               (*
               FOR #Temp_Index_i := #ServerVersion_StartNum TO #MessageLen - 1 DO   //去掉前面的8个数据，同时从0开始，所以-9
                   #SaltString[#Temp_Index_i - #ServerVersion_StartNum + 2] := #REV_Buffer[#ServerVersion_StartNum];//挑战字符串的后面N个Byte
                   #ServerVersion_StartNum := #ServerVersion_StartNum + 1;
               END_FOR;*)
           END_REGION

           REGION Client_Auth_Packet
               #Temp_NowNum := 0;
               #Client_MaxLen := DINT_TO_DWORD(#MessageMaxLen);
               // Length                            3     Byte   最后处理
               #Temp_NowNum := #Temp_NowNum +3;
               // Sequence                      1     Byte
               #SND_Buffer[#Temp_NowNum] :=SINT_TO_BYTE( DINT_TO_SINT(#CDD.Connect_Sequence + 1));
               #Temp_NowNum := #Temp_NowNum + 1;
               // CapabilityFlag               4     Byte
               #SND_Buffer[#Temp_NowNum] := #Client_CapabilityFlag.%B0;
               #Temp_NowNum := #Temp_NowNum + 1;
               #SND_Buffer[#Temp_NowNum] := #Client_CapabilityFlag.%B1;
               #Temp_NowNum := #Temp_NowNum + 1;
               #SND_Buffer[#Temp_NowNum] := #Client_CapabilityFlag.%B2;
               #Temp_NowNum := #Temp_NowNum + 1;
               #SND_Buffer[#Temp_NowNum] := #Client_CapabilityFlag.%B3;
               #Temp_NowNum := #Temp_NowNum + 1;
               // Max_Length                   4     Byte
               #SND_Buffer[#Temp_NowNum] := #Client_MaxLen.%B0;
               #Temp_NowNum := #Temp_NowNum + 1;
               #SND_Buffer[#Temp_NowNum] := #Client_MaxLen.%B1;
               #Temp_NowNum := #Temp_NowNum + 1;
               #SND_Buffer[#Temp_NowNum] := #Client_MaxLen.%B2;
               #Temp_NowNum := #Temp_NowNum + 1;
               #SND_Buffer[#Temp_NowNum] := #Client_MaxLen.%B3;
               #Temp_NowNum := #Temp_NowNum + 1;
               // CharacterSet                 1     Byte
               #SND_Buffer[#Temp_NowNum] := #CDD.Server_Character_Set;
               #Temp_NowNum := #Temp_NowNum + 1;
               // Fill Data  (16#00)          23  Byte
               FOR #Temp_Index_i := 0 TO 22 DO
                   #SND_Buffer[#Temp_NowNum + #Temp_Index_i] := b#16#00;
               END_FOR;
               #Temp_NowNum := #Temp_NowNum + 23;
               // User Name                    N    Byte    Last Character    16#00
               #Temp_StrLen := LEN(#UserName);
               FOR #Temp_Index_i := 0 TO #Temp_StrLen - 1 DO
                   #SND_Buffer[#Temp_NowNum + #Temp_Index_i] := #UserName[#Temp_Index_i + 1];
               END_FOR;
               #Temp_NowNum := #Temp_NowNum + #Temp_StrLen;
               #SND_Buffer[#Temp_NowNum] := b#16#00;
               #Temp_NowNum := #Temp_NowNum + 1;
               #SND_Buffer[#Temp_NowNum] := b#16#14;
               #Temp_NowNum := #Temp_NowNum + 1;
               // Token                              N    Byte    Last Character    16#00
               #Calc_Encryption_SHA1(IN_Str := #PassWord,
                                     TempOutStr => #Temp_SHA1);
               #Calc_Encryption_SHA1(IN_Str := #Temp_SHA1,
                                     Len:=20,
                                     TempOutStr => #Temp_SHA1_2);
               // Strg_TO_Chars(Strg := #PassWord,
               //               pChars := 0,
               //               Cnt => #Temp_SHA_Arry_Num,
               //               Chars := #Temp_SHA_Arry);
               // #Temp_SHA_Arry_Num_Int := UINT_TO_INT(#Temp_SHA_Arry_Num);

               FOR #Temp_Index_i := 0 TO 19 DO
                   #Temp_SHA_Arry[#Temp_Index_i] := #SaltString[#Temp_Index_i];
               END_FOR;
               FOR #Temp_Index_i := 20 TO 39 DO
                   #Temp_SHA_Arry[#Temp_Index_i] := #Temp_SHA1_2[#Temp_Index_i - 20];
               END_FOR;

               #Calc_Encryption_SHA1(IN_Str := #Temp_SHA_Arry,
                                     Len := 40,
                                     TempOutStr => #Temp_SHA1_3);

               FOR #Temp_Index_i := 0 TO 19 DO
                   #Token[#Temp_Index_i] := #Temp_SHA1[#Temp_Index_i] XOR #Temp_SHA1_3[#Temp_Index_i];
                   #SND_Buffer[#Temp_NowNum + #Temp_Index_i] := #Token[#Temp_Index_i];
               END_FOR;
               #Temp_NowNum := #Temp_NowNum + 20;
               #SND_Buffer[#Temp_NowNum] := b#16#00;
               #Temp_NowNum := #Temp_NowNum + 1;

               // DataBase Name           N    Byte    Last Character    16#00
               #Temp_StrLen := LEN(#DB_Name);
               FOR #Temp_Index_i := 0 TO #Temp_StrLen - 1 DO
                   #SND_Buffer[#Temp_NowNum + #Temp_Index_i] := #DB_Name[#Temp_Index_i + 1];
               END_FOR;
               #Temp_NowNum := #Temp_NowNum + #Temp_StrLen;
               #SND_Buffer[#Temp_NowNum] := b#16#00;
               #Temp_NowNum := #Temp_NowNum + 1;
               //CLIENT_PLUGIN_AUTH
               #Temp_StrLen := LEN(#CDD.CLIENT_PLUGIN_AUTH);
               FOR #Temp_Index_i := 0 TO #Temp_StrLen - 1 DO
                   #SND_Buffer[#Temp_NowNum + #Temp_Index_i] := #CDD.CLIENT_PLUGIN_AUTH[#Temp_Index_i + 1];
               END_FOR;
               #Temp_NowNum := #Temp_NowNum + #Temp_StrLen;
               #SND_Buffer[#Temp_NowNum] := b#16#00;
               #Temp_NowNum := #Temp_NowNum + 1;

               //数据长度写入前三个byte
               #Temp_Dword := DINT_TO_DWORD(INT_TO_DINT(#Temp_NowNum - 4));
               #SND_Buffer[0] := #Temp_Dword.%B0;
               #SND_Buffer[1] := #Temp_Dword.%B1;
               #SND_Buffer[2] := #Temp_Dword.%B2;
               #Step := 3;
               #NetSendLen := #Temp_NowNum;
           END_REGION

           ;

       3:  // 等待发送完成
           #NetRcv_EN := TRUE;
           #NetSend_EN := TRUE;
           IF #NetSend_Done THEN
               #NetSend_Done := FALSE;
               #NetSend_EN := FALSE;
               #Step := 4;
           END_IF;

       4:  // 等待接收数据

           IF    #NetRcv_Done  THEN
               #NetRcv_Done := FALSE;

              // #NetRcv_Len := UDINT_TO_INT(#NetRcv.RCVD_LEN);
               #NetRcv_EN := FALSE;
               #Step := 5;
           END_IF;
       5:  // 如果在等待服务器第一次连接
           IF #REV_Buffer[5]=b#16#00 AND  #NetRcv_Len >7 THEN
               #Temp_CND := TRUE;
               #NetRcv_EN := TRUE;
           END_IF;


       6:  // 申请服务器断开连接
            #SND_Buffer[0] := b#16#01;
            #SND_Buffer[1] := b#16#00;
            #SND_Buffer[2] := b#16#00;
            #SND_Buffer[3] := b#16#00;
            #SND_Buffer[4] := b#16#01;
            #NetSendEnd_EN := TRUE;
            IF #NetSendEnd_Done THEN
                #Step := 7;
            END_IF;

        7:  // 申请服务器断开连接

            #NetDiscon_EN := TRUE;
        8:
            ;
       ELSE  // Statement section ELSE
           ;
   END_CASE;


   (***********************************************************发送数据******************************************************************)
       #NetSend(REQ := #NetSend_EN,
                ID := #Net_ID,
                // DONE=>#NetSend_Done,
                LEN := INT_TO_UDINT(#NetSendLen),// INT_TO_UINT(#Temp_NowNum),
                DATA := #SND_Buffer);
       IF #NetSend.DONE THEN
           #NetSend_Done := TRUE;
       END_IF;

       #NetSendEnd(REQ := #NetSendEnd_EN,
                   ID := #Net_ID,
                   LEN := 5,
                   DONE => #NetSendEnd_Done,
                   DATA := #SND_Buffer);





   (***********************************************************断开连接******************************************************************)

   #NetDISCON(REQ:=#NetDiscon_EN AND #Timer_ON.Q ,
              ID:=#Net_ID);

   #Timer_ON(IN := NOT #Timer_OFF.Q,
             PT := t#0.5s);

   #Timer_OFF(IN := #Timer_ON.Q,
              PT := t#0.5s);




   (***********************************************************监测连接******************************************************************)
   #NetDiag(REQ := #Timer_ON.Q,
            ID := #Net_ID,
            RESULT := #TDiag_Result);
   IF  #NetDiag.ERROR THEN
       #Temp_ConnStatus := B#16#00;
   END_IF;
   IF #NetDiag.DONE THEN
       #Temp_ConnStatus := #TDiag_Result.State;
   END_IF;
   IF #Temp_ConnStatus <> B#16#04 THEN
       #Temp_CND := FALSE;
   END_IF;

   #CDD.Connect_OK := #Temp_CND;

   #Timer_Error(IN := #Connect AND NOT #Temp_CND,
                PT := t#10s);

   #Error := #Timer_Error.Q;
   #CND := #Temp_CND;
   #ConnStatus := #Temp_ConnStatus;

   (***********************************************************数据传递******************************************************************)
   #CDD.Recv_Buffer := #REV_Buffer;
   IF #NetRcv.NDR THEN
       #CDD.Recv_Done := TRUE;
       #CDD.Recv_Len := UDINT_TO_INT(#NetRcv.RCVD_LEN);
   END_IF;
END_FUNCTION_BLOCK

FUNCTION_BLOCK "uMySQL_Query"   // FB5, SCL
{ S7_Optimized_Access := 'TRUE' }
VERSION : 0.1
   VAR_INPUT
      Command : WString[2048];
      Execute : Bool;
   END_VAR
   VAR_OUTPUT
      Done : Bool;
      Busy : Bool;
      Error : Bool;
   END_VAR
   VAR_IN_OUT
      CDD : "uMySQL_CDD";
   END_VAR
   VAR
      Net_Send : TSEND;
      Net_Send_EN : Bool;
      Net_Send_Done : Bool;
      Net_Send_Len : UInt;
      Command_Len : UInt;
      Net_Recv_EN : Bool;
      Net_Recv_Done : Bool;
      Net_Recv_Len : UInt;
      Temp_Bool : Array[0..19] of Bool;
      SendBuffer : Array[0..2048] of Byte;
      RecvBuffer : Array[0..2048] of Byte;
      SendBufferWChar : Array[0..2048] of WChar;
      TRCV : TRCV;
      Function_Run : Bool;
      Timer_instance : TON_TIME;
   END_VAR
   VAR_TEMP
      Temp_Index_i : Int;
      Temp_Dword : DWord;
      Temp_word : Word;
      Temp_Num : Int;
   END_VAR
BEGIN

   IF #Execute THEN
       #Function_Run:= TRUE;
   END_IF;

   IF #Function_Run AND NOT #Temp_Bool[0] THEN
       #Temp_Bool[0] := TRUE;
       #Net_Send_EN := TRUE;
       #Command_Len := INT_TO_UINT(LEN(#Command));
       #SendBuffer[4] := B#16#03;

       Strg_TO_Chars(Strg := #Command,
                     pChars := 0,
                     Cnt => #Command_Len,
                     Chars := #SendBufferWChar);
       (*  
       FOR #Temp_Index_i := 0 TO UINT_TO_INT( #Command_Len) -1 DO
           #SendBuffer[#Temp_Index_i + 5]:=WCHAR_TO_BYTE(#SendBufferWChar[#Temp_Index_i]) ;

       END_FOR;
       #Net_Send_Len := #Command_Len + 5;
       *)
       #Net_Send_Len := 5;

       FOR #Temp_Index_i := 0 TO UINT_TO_INT(#Command_Len) - 1 DO

           #Temp_Dword := "Wchar_To_UTF8"("WChar" := #SendBufferWChar[#Temp_Index_i], Num => #Temp_Num);
           CASE #Temp_Num OF
               1:  // 如果是单字符
                   #SendBuffer[#Net_Send_Len] := #Temp_Dword.%B0;
                   #Net_Send_Len := #Net_Send_Len + 1;
               2:  // 如果是两字节
                   #SendBuffer[#Net_Send_Len] := #Temp_Dword.%B1;
                   #Net_Send_Len := #Net_Send_Len + 1;
                   #SendBuffer[#Net_Send_Len] := #Temp_Dword.%B0;
                   #Net_Send_Len := #Net_Send_Len + 1;
               ELSE  // 如果是其他情况
                   #SendBuffer[#Net_Send_Len] := #Temp_Dword.%B2;
                   #Net_Send_Len := #Net_Send_Len + 1;
                   #SendBuffer[#Net_Send_Len] := #Temp_Dword.%B1;
                   #Net_Send_Len := #Net_Send_Len + 1;
                   #SendBuffer[#Net_Send_Len] := #Temp_Dword.%B0;
                   #Net_Send_Len := #Net_Send_Len + 1;
           END_CASE;

       END_FOR;

       #Net_Send_EN := TRUE; 
                                 //数据长度写入前三个byte
                                 #Temp_Dword := DINT_TO_DWORD(INT_TO_DINT(UINT_TO_INT(#Net_Send_Len) - 4));
                                 #SendBuffer[0] := #Temp_Dword.%B0;
                                 #SendBuffer[1] := #Temp_Dword.%B1;
                                 #SendBuffer[2] := #Temp_Dword.%B2;
                             END_IF;


   IF NOT #Function_Run THEN
       #Temp_Bool[0] := FALSE;
       #Net_Recv_Len := 0;
       #Net_Recv_Done := FALSE;
       #Net_Send_EN := FALSE;
       #Net_Recv_EN := FALSE;
       #Error := FALSE;
       #Done := FALSE;
   END_IF;


   #Net_Send(REQ:=#Net_Send_EN,
             ID:=#CDD.Connect_ID,
             LEN:=#Net_Send_Len,
             DONE=>#Net_Send_Done,
             DATA:=#SendBuffer);

   IF #Net_Send.DONE OR #Net_Send.ERROR THEN
       #Net_Send_EN := FALSE;
       #Function_Run := FALSE;
       IF #Net_Send.ERROR THEN
           #Error := TRUE;
       END_IF;
   END_IF;


   IF #CDD.Recv_Done AND #Function_Run THEN
       #Temp_word.%B0 := #CDD.Recv_Buffer[0];
       #Temp_word.%B1 := #CDD.Recv_Buffer[1];
       IF #CDD.Recv_Len = (WORD_TO_INT(#Temp_word)+4) THEN

           CASE BYTE_TO_INT(#CDD.Recv_Buffer[4]) OF
               0:
                   #Done := TRUE;
               255:  // Statement section case 2 to 4
                   #Error := TRUE;
               ELSE  // Statement section ELSE
                   ;
           END_CASE; //通过返回的数据判断是否执行成功
       ELSE
           #Error := TRUE;//如果接收的数据长度和范围数据中给定的不同则认定是通信错误
       END_IF;
       #CDD.Recv_Done := FALSE;
   END_IF;


   #Timer_instance(IN:=#Function_Run AND ( NOT #Done),
                   PT:=t#1s  );
   IF #Timer_instance.Q THEN    //如果命令执行超时，也认为是故障
       #Error := TRUE;
   END_IF;

   IF #Error THEN
       #Function_Run := FALSE;
   END_IF;
   IF #Done THEN
       #Function_Run := FALSE;
   END_IF;
END_FUNCTION_BLOCK

FUNCTION_BLOCK "Calc_Encryption_SHA1"   // FB6, SCL
{ S7_Optimized_Access := 'FALSE' }
VERSION : 0.1
   VAR_INPUT
      IN_Str : Variant;
      Len : Int;
   END_VAR
   VAR_OUTPUT
      TempOutStr : Array[0..19] of Byte;
      Encrption AT TempOutStr : Array[0..4] of DWord;
   END_VAR
   VAR_TEMP
      "A" : DWord;
      "B" : DWord;
      C : DWord;
      D : DWord;
      "E" : DWord;
      Length : Int;
      Lenth_Uint : UInt;
      MessageBlock : Array[0..63] of Byte;
      MessageBlock_DWORD AT MessageBlock : Array[0..15] of DWord;
      W : Array[0..79] of DWord;
      Index_i : Int;
      temp : DWord;
      Temp_Str : String;
      Temp_Array : Array[0..446] of Byte;
   END_VAR
   VAR CONSTANT
      K0 : DWord := 16#5A827999;   // K0计算常量
      K1 : DWord := 16#6ED9EBA1;   // K1计算常量
      K2 : DWord := 16#8F1BBCDC;   // K2计算常量
      K3 : DWord := 16#CA62C1D6;   // K3计算常量
      Const_A : DWord := 16#67452301;   // 链接变量A
      Const_B : DWord := 16#EFCDAB89;   // 链接变量B
      Const_C : DWord := 16#98BADCFE;   // 链接变量C
      Const_D : DWord := 16#10325476;   // 链接变量D
      Const_E : DWord := 16#C3D2E1F0;   // 链接变量E
   END_VAR
BEGIN
   (***************************************************数据初始化******************************************************)
   #A := #Const_A;
   #B := #Const_B;
   #C := #Const_C;
   #D := #Const_D;
   #E := #Const_E;
   //#Length := LEN(#IN_Str);
   FILL_BLK(IN := B#16#00,  COUNT := 64,  OUT => #MessageBlock[0]);
   FILL_BLK(IN := DW#16#000000000,   COUNT := 80,  OUT => #W[0]);




   (*************************************************填充/准备数据****************************************************)
   IF TypeOf(#IN_Str) =String THEN
       //如果是字符串
       VariantGet(SRC:=#IN_Str,
                  DST=>#Temp_Str);
       #Length := LEN(#Temp_Str);

       Strg_TO_Chars(Strg :=#Temp_Str ,
                     pChars := 0,
                     Cnt => #Lenth_Uint,
                     Chars := #MessageBlock);   //填充客户输入字符
   ELSE
       IF IS_ARRAY(#IN_Str) THEN
          // #Length:=UDINT_TO_INT(CountOfElements(#IN_Str)) ;
           #Length := #Len;
           VariantGet(SRC:=#IN_Str,     DST=>#Temp_Array);
           MOVE_BLK(IN := #Temp_Array[0],  COUNT :=INT_TO_UINT( #Length),  OUT => #MessageBlock[0]);
       END_IF;
     ;
   END_IF;
   (*********************************************输入数据安全检测****************************************************)
   IF (#Length = 0) OR (#Length > 56) THEN
       RETURN;
   END_IF;

   #MessageBlock[#Length] := B#16#80;   //后一位填1，其他全为0
   #MessageBlock_DWORD[14] :=DW#16#00000000;          //填充数据长度高位
   #MessageBlock_DWORD[15] := DINT_TO_DWORD(#Length * 8);//填充数据长度低位
   MOVE_BLK(IN := #MessageBlock_DWORD[0],  COUNT := 16,  OUT => #W[0]);
   FOR #Index_i := 16 TO 79 DO
       #W[#Index_i] := ROL(N := 1, IN := (#W[#Index_i - 3] XOR #W[#Index_i - 8] XOR #W[#Index_i - 14] XOR #W[#Index_i - 16]));
   END_FOR;
   (*************************************************计算过程****************************************************)
   FOR #Index_i := 0 TO 19 DO
       #temp := ROL(IN := #A, N := 5) + ((#B AND #C) OR (NOT (#B) AND #D)) + #E + #W[#Index_i] + #K0;
       #E := #D;
       #D := #C;
       #C := ROL(IN := #B, N := 30);
       #B := #A;
       #A := #temp;
   END_FOR;

   FOR #Index_i := 20 TO 39 DO
       #temp := ROL(IN := #A, N := 5) + (#B XOR #C XOR #D) + #E + #W[#Index_i] + #K1;
       #E := #D;
       #D := #C;
       #C := ROL(N := 30, IN := #B);
       #B := #A;
       #A := #temp;
   END_FOR;

   FOR #Index_i := 40 TO 59 DO
       #temp := ROL(N := 5, IN := #A) + ((#B AND #C) OR (#B AND #D) OR (#C AND #D)) + #E + #W[#Index_i] + #K2;
       #E := #D;
       #D := #C;
       #C := ROL(N := 30, IN := #B);
       #B := #A;
       #A := #temp;
   END_FOR;

   FOR #Index_i := 60 TO 79 DO
       #temp := ROL(N := 5, IN := #A) + (#B XOR #C XOR #D) + #E + #W[#Index_i] + #K3;
       #E := #D;
       #D := #C;
       #C := ROL(N := 30, IN := #B);
       #B := #A;
       #A := #temp;
   END_FOR;

   #Encrption[0] := #Const_A + #A;
   #Encrption[1] := #Const_B+ #B;
   #Encrption[2] := #Const_C + #C;
   #Encrption[3] := #Const_D + #D;
   #Encrption[4] := #Const_E + #E;
END_FUNCTION_BLOCK

FUNCTION_BLOCK "uMySQL_Use"   // FB8, SCL
{ S7_Optimized_Access := 'TRUE' }
VERSION : 0.1
   VAR_INPUT
      DB_Name : WString[2048];
      Execute : Bool;
   END_VAR
   VAR_OUTPUT
      Done : Bool;
      Busy : Bool;
      Error : Bool;
   END_VAR
   VAR_IN_OUT
      CDD : "uMySQL_CDD";
   END_VAR
   VAR
      Net_Send : TSEND;
      Net_Send_EN : Bool;
      Net_Send_Done : Bool;
      Net_Send_Len : UInt;
      Command_Len : UInt;
      Net_Recv_EN : Bool;
      Net_Recv_Done : Bool;
      Net_Recv_Len : UInt;
      Temp_Bool : Array[0..19] of Bool;
      SendBuffer : Array[0..2048] of Byte;
      RecvBuffer : Array[0..2048] of Byte;
      SendBufferWChar : Array[0..2048] of WChar;
      TRCV : TRCV;
      Function_Run : Bool;
      Timer_instance : TON_TIME;
   END_VAR
   VAR_TEMP
      Temp_Index_i : Int;
      Temp_Dword : DWord;
      Temp_word : Word;
   END_VAR
BEGIN

   IF #Execute THEN
       #Function_Run:= TRUE;
   END_IF;

   IF #Function_Run AND NOT #Temp_Bool[0] THEN
       #Temp_Bool[0] := TRUE;
       #Net_Send_EN := TRUE;
       #Command_Len := INT_TO_UINT(LEN(#DB_Name));
       #SendBuffer[4] := B#16#02;

       Strg_TO_Chars(Strg := #DB_Name,
                     pChars := 0,
                     Cnt => #Command_Len,
                     Chars := #SendBufferWChar);

       FOR #Temp_Index_i := 0 TO UINT_TO_INT(#Command_Len) - 1 DO
           #SendBuffer[#Temp_Index_i + 5] := WCHAR_TO_BYTE(#SendBufferWChar[#Temp_Index_i]);
       END_FOR;
       #Net_Send_Len := #Command_Len + 5;
       #Net_Send_EN := TRUE;
       //数据长度写入前三个byte
       #Temp_Dword := DINT_TO_DWORD(INT_TO_DINT(UINT_TO_INT(#Net_Send_Len) - 4));
       #SendBuffer[0] := #Temp_Dword.%B0;
       #SendBuffer[1] := #Temp_Dword.%B1;
       #SendBuffer[2] := #Temp_Dword.%B2;
   END_IF;


   IF NOT #Function_Run THEN
       #Temp_Bool[0] := FALSE;
       #Net_Recv_Len := 0;
       #Net_Recv_Done := FALSE;
       #Net_Send_EN := FALSE;
       #Net_Recv_EN := FALSE;
       #Error := FALSE;
       #Done := FALSE;
   END_IF;


   #Net_Send(REQ:=#Net_Send_EN,
             ID:=#CDD.Connect_ID,
             LEN:=#Net_Send_Len,
             DONE=>#Net_Send_Done,
             DATA:=#SendBuffer);

   IF #Net_Send.DONE OR #Net_Send.ERROR THEN
       #Net_Send_EN := FALSE;
       #Function_Run := FALSE;
       IF #Net_Send.ERROR THEN
           #Error := TRUE;
       END_IF;
   END_IF;


   IF #CDD.Recv_Done AND #Function_Run THEN
       #Temp_word.%B0 := #CDD.Recv_Buffer[0];
       #Temp_word.%B1 := #CDD.Recv_Buffer[1];
       IF #CDD.Recv_Len = (WORD_TO_INT(#Temp_word)+4) THEN

           CASE BYTE_TO_INT(#CDD.Recv_Buffer[4]) OF
               0:
                   #Done := TRUE;
               255:  // Statement section case 2 to 4
                   #Error := TRUE;
               ELSE  // Statement section ELSE
                   ;
           END_CASE; //通过返回的数据判断是否执行成功
       ELSE
           #Error := TRUE;//如果接收的数据长度和范围数据中给定的不同则认定是通信错误
       END_IF;
       #CDD.Recv_Done := FALSE;
   END_IF;

   #Timer_instance(IN:=#Function_Run AND ( NOT #Done),
                   PT:=t#1s  );
   IF #Timer_instance.Q THEN    //如果命令执行超时，也认为是故障
       #Error := TRUE;
   END_IF;

   IF #Error THEN
       #Function_Run := FALSE;
   END_IF;
   IF #Done THEN
       #Function_Run := FALSE;
   END_IF;
END_FUNCTION_BLOCK

FUNCTION_BLOCK "uMySQL_Command"   // FB909, SCL
{ S7_Optimized_Access := 'TRUE' }
VERSION : 0.1
   VAR
      Command : WString[2048];
   END_VAR
   VAR_TEMP
      TempStr : WString;
   END_VAR
BEGIN
   "数据库字符串"."wstring" :=WSTRING#'INSERT INTO rb001011(Addr,temp_LF,temp_RF,temp_LB,temp_RB,Distance_L,Distance_R,';
   "数据库字符串"."wstring" := CONCAT(IN1 := "数据库字符串"."wstring", IN2 := WSTRING#'Motor_Current,Motor_Freq,Motor_Power,Motor_Eng,Motor_Runhours,');
   "数据库字符串"."wstring" := CONCAT(IN1 := "数据库字符串"."wstring", IN2 := WSTRING#'EN_Temp,EN_RH,temp_Ruber,');
   "数据库字符串"."wstring" := CONCAT(IN1 := "数据库字符串"."wstring", IN2 := WSTRING#'Motor_Ready,Motor_Running,Motor_Fault,');
   "数据库字符串"."wstring" := CONCAT(IN1 := "数据库字符串"."wstring", IN2 := WSTRING#'SerialNum,Operator');
   "数据库字符串"."wstring" := CONCAT(IN1 := "数据库字符串"."wstring", IN2 := WSTRING#')VALUES(');

   "数据库字符串"."wstring" := CONCAT(IN1 := "数据库字符串"."wstring", IN2 := "uMySQL_Aux_ConnectValue"(Value := "数据库字符串".Addr,
                                                                                                                         PREC := 3,
                                                                                                                         Tail := WSTRING#','));
   "数据库字符串"."wstring" := CONCAT(IN1 := "数据库字符串"."wstring", IN2 := "uMySQL_Aux_ConnectValue"(Value := "数据库字符串".UploadData.左前辊温度,
                                                                                                                         PREC := 3,
                                                                                                                         Tail := WSTRING#','));

   "数据库字符串"."wstring" := CONCAT(IN1 := "数据库字符串"."wstring", IN2 := "uMySQL_Aux_ConnectValue"(Value :="数据库字符串".UploadData.右前辊温度,
                                                                                                                         PREC := 3,
                                                                                                                         Tail := WSTRING#','));
   "数据库字符串"."wstring" := CONCAT(IN1 := "数据库字符串"."wstring", IN2 := "uMySQL_Aux_ConnectValue"(Value := "数据库字符串".UploadData.左后辊温度,
                                                                                                                         PREC := 3,
                                                                                                                         Tail := WSTRING#','));
   "数据库字符串"."wstring" := CONCAT(IN1 := "数据库字符串"."wstring", IN2 := "uMySQL_Aux_ConnectValue"(Value := "数据库字符串".UploadData.右后辊温度,
                                                                                                                         PREC := 3,
                                                                                                                         Tail := WSTRING#','));
   "数据库字符串"."wstring" := CONCAT(IN1 := "数据库字符串"."wstring", IN2 := "uMySQL_Aux_ConnectValue"(Value := "数据库字符串".UploadData.左间隙,
                                                                                                                         PREC := 3,
                                                                                                                         Tail := WSTRING#','));


   "数据库字符串"."wstring" := CONCAT(IN1 := "数据库字符串"."wstring", IN2 := "uMySQL_Aux_ConnectValue"(Value := "数据库字符串".UploadData.右间隙,
                                                                                                                         PREC := 3,
                                                                                                                         Tail := WSTRING#','));
   "数据库字符串"."wstring" := CONCAT(IN1 := "数据库字符串"."wstring", IN2 := "uMySQL_Aux_ConnectValue"(Value := "数据库字符串".UploadData.滚筒电机电流,
                                                                                                                         PREC := 3,
                                                                                                                         Tail := WSTRING#','));
   "数据库字符串"."wstring" := CONCAT(IN1 := "数据库字符串"."wstring", IN2 := "uMySQL_Aux_ConnectValue"(Value := "数据库字符串".UploadData.滚筒电机频率,
                                                                                                                         PREC := 3,
                                                                                                                         Tail := WSTRING#','));
   "数据库字符串"."wstring" := CONCAT(IN1 := "数据库字符串"."wstring", IN2 := "uMySQL_Aux_ConnectValue"(Value := "数据库字符串".UploadData.滚筒电机功率,
                                                                                                                         PREC := 3,
                                                                                                                         Tail := WSTRING#','));
   "数据库字符串"."wstring" := CONCAT(IN1 := "数据库字符串"."wstring", IN2 := "uMySQL_Aux_ConnectValue"(Value := "数据库字符串".UploadData.滚筒电机电度,
                                                                                                                         PREC := 3,
                                                                                                                         Tail := WSTRING#','));
   "数据库字符串"."wstring" := CONCAT(IN1 := "数据库字符串"."wstring", IN2 := "uMySQL_Aux_ConnectValue"(Value := "数据库字符串".UploadData.滚筒电机计时,
                                                                                                                         PREC := 3,
                                                                                                                         Tail := WSTRING#','));



   "数据库字符串"."wstring" := CONCAT(IN1 := "数据库字符串"."wstring", IN2 := "uMySQL_Aux_ConnectValue"(Value := "数据库字符串".UploadData.环境温度,
                                                                                                                         PREC := 3,
                                                                                                                         Tail := WSTRING#','));

   "数据库字符串"."wstring" := CONCAT(IN1 := "数据库字符串"."wstring", IN2 := "uMySQL_Aux_ConnectValue"(Value := "数据库字符串".UploadData.环境湿度,
                                                                                                                         PREC := 3,
                                                                                                                         Tail := WSTRING#','));

   "数据库字符串"."wstring" := CONCAT(IN1 := "数据库字符串"."wstring", IN2 := "uMySQL_Aux_ConnectValue"(Value := "数据库字符串".UploadData.胶温,
                                                                                                                         PREC := 3,
                                                                                                                         Tail := WSTRING#','));




   "数据库字符串"."wstring" := CONCAT(IN1 := "数据库字符串"."wstring", IN2 := "uMySQL_Aux_ConnectValue"(Value := "数据库字符串".UploadData.开关量汇总.%X0,
                                                                                                                         PREC := 1,
                                                                                                                         Tail := WSTRING#','));


   "数据库字符串"."wstring" := CONCAT(IN1 := "数据库字符串"."wstring", IN2 := "uMySQL_Aux_ConnectValue"(Value := "数据库字符串".UploadData.开关量汇总.%X1,
                                                                                                                         PREC := 1,
                                                                                                                         Tail := WSTRING#','));

   "数据库字符串"."wstring" := CONCAT(IN1 := "数据库字符串"."wstring", IN2 := "uMySQL_Aux_ConnectValue"(Value := "数据库字符串".UploadData.开关量汇总.%X2,
                                                                                                                         PREC := 1,
                                                                                                                         Tail := WSTRING#','));
   "数据库字符串"."wstring" := CONCAT(IN1 := "数据库字符串"."wstring", IN2 := "uMySQL_Aux_ConnectValue"(Value :="数据库字符串".UploadData.当前任务编号,
                                                                                                                         PREC := 1,
                                                                                                                         Tail := WSTRING#','));
   "数据库字符串"."wstring" := CONCAT(IN1 := "数据库字符串"."wstring", IN2 := "uMySQL_Aux_ConnectValue"(Value := "数据库字符串".UploadData.当前人员编号,
                                                                                                                         PREC := 1,
                                                                                                                         Tail := WSTRING#')'));
END_FUNCTION_BLOCK

FUNCTION "uMySQL_Aux_ConnectValue" : WString   // FC160, SCL
{ S7_Optimized_Access := 'TRUE' }
VERSION : 0.1
   VAR_INPUT
      Value : Variant;
      PREC : USInt;
      Tail : WString;
   END_VAR
   VAR_TEMP
      Value_Real : Real;
      Value_Int : Int;
      Value_Dint : DInt;
      Value_Bool : Bool;
      Value_Wstring : WString;
      Temp_Str : WString[2048];
      Temp_Command : WString[2048];
      Value_M : Int;
      Value_FP : USInt;
      Value_PP : USInt;
      Valve_Format : Word;
      TempWstring_Len : Int;
      TempWstring_Index : Int;
   END_VAR
BEGIN
   #Value_Bool:=FALSE;
   #Value_Real := 0.0;
   #Temp_Command:=WSTRING#'';
   IF TypeOf(#Value_Bool) = TypeOf(#Value) THEN
       VariantGet(SRC := #Value,
                  DST => #Value_Bool);
       IF #Value_Bool THEN
           #Temp_Command := WSTRING#'1';
       ELSE
           #Temp_Command := WSTRING#'0';
       END_IF;
   ELSIF TypeOf(#Value_Wstring) = TypeOf(#Value) THEN //开始处理字符串
       VariantGet(SRC := #Value,
                  DST => #Value_Wstring);
       #TempWstring_Len := LEN(#Value_Wstring);
       #Temp_Command := CONCAT(IN1 := wstring#'"', IN2 := #Value_Wstring);
       // FOR #TempWstring_Index := 1 TO #TempWstring_Len DO

       //     IF _condition_ THEN
       //         // Statement section IF
       //         ;
       //     END_IF;

       //     ;
       // END_FOR;

       #Temp_Command := CONCAT(IN1 := #Temp_Command, IN2 := wstring#'"'); //字符串处理结束

   ELSE


       IF TypeOf(#Value_Int) = TypeOf(#Value) THEN
           VariantGet(SRC := #Value,
                      DST => #Value_Int);
           #Value_Real := INT_TO_REAL(#Value_Int);
           #Value_FP := 0;
           #Value_PP := 0;
       ELSIF TypeOf(#Value_Dint) = TypeOf(#Value) THEN
           VariantGet(SRC := #Value,
                      DST => #Value_Dint);
           #Value_Real := DINT_TO_REAL(#Value_Dint);
           #Value_FP := 0;
           #Value_PP := 0;

       ELSE
           VariantGet(SRC := #Value,
                      DST => #Value_Real);
           #Value_FP := #PREC;
           #Value_PP := 1;
       END_IF;

       #Valve_Format := 16#0000;
       IF #Value_Real < 0.0 THEN
           #Valve_Format := 16#0004;
           #Value_PP := #Value_PP + 2;
       END_IF;
       #Value_M := #Value_FP + 1;
       IF ABS(#Value_Real / 10) >= 1 THEN
           #Value_M := #Value_FP + 2;
       END_IF;
       IF ABS(#Value_Real / 100) >= 1 THEN
           #Value_M := #Value_FP + 3;
       END_IF;

       IF ABS(#Value_Real / 1000) >= 1 THEN
           #Value_M := #Value_FP + 4;
       END_IF;

       IF ABS(#Value_Real / 10000) >= 1 THEN
           #Value_M := #Value_FP + 5;
       END_IF;

       IF ABS(#Value_Real / 100000) >= 1 THEN
           #Value_M := #Value_FP + 6;
       END_IF;
       IF ABS(#Value_Real / 1000000) >= 1 THEN
           #Value_M := #Value_FP + 7;
       END_IF;
       IF ABS(#Value_Real / 10000000) >= 1 THEN
           #Value_M := #Value_FP + 8;
       END_IF;
       IF ABS(#Value_Real / 100000000) >= 1 THEN
           #Value_M := #Value_FP + 9;
       END_IF;
       IF ABS(#Value_Real / 1000000000) >= 1 THEN
           #Value_M := #Value_FP + 10;
       END_IF;

       IF TypeOf(#Value_Dint) = TypeOf(#Value) THEN
           VAL_STRG(IN := #Value_Dint,
                    SIZE := INT_TO_USINT(#Value_M) + #Value_PP,
                    PREC := #Value_FP,
                    FORMAT := #Valve_Format,
                    P := 1,
                    OUT => #Temp_Command);
       ELSE
           VAL_STRG(IN := #Value_Real,
                    SIZE := INT_TO_USINT(#Value_M) + #Value_PP,
                    PREC := #Value_FP,
                    FORMAT := #Valve_Format,
                    P := 1,
                    OUT => #Temp_Command);
       END_IF;




   END_IF;





   #Temp_Str:= CONCAT(IN1 := wstring#'', IN2 := #Temp_Command);
   //#Temp_Str := "LWString_Connect"(S1 := #CommandLine, S2 := #Temp_Command);


   #Temp_Str := CONCAT(IN1 := #Temp_Str, IN2 := #Tail);
   //#Temp_Str := "LWString_Connect"(S1 := #Temp_Str, S2 :=  #Tail);
   #uMySQL_Aux_ConnectValue := #Temp_Str;
END_FUNCTION

FUNCTION "LWString_Connect" : WString   // FC161, LAD
{ S7_Optimized_Access := 'TRUE' }
VERSION : 0.1
   VAR_INPUT
      S1 : WString;
      S2 : WString;
   END_VAR
   VAR_TEMP
      Array_S1 : Array[0..2048] of WChar;
      Array_S2 : Array[0..4096] of WChar;
      LEN_S1 : UInt;
      LEN_S2 : UInt;
      LEN : UInt;
   END_VAR
BEGIN

REGION Network 1
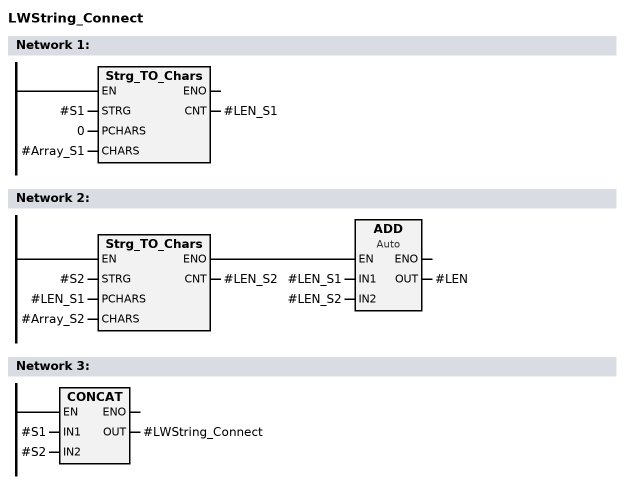
   // no SCL statement known for Strg_TO_Chars: written as a call
   Strg_TO_Chars(Strg := #S1, pChars := 0, Chars := #Array_S1, Cnt => #LEN_S1);
END_REGION

REGION Network 2
   // no SCL statement known for Strg_TO_Chars: written as a call
   // ENO of a box is taken as its EN; it also drops when the box reports an error
   Strg_TO_Chars(Strg := #S2, pChars := #LEN_S1, Chars := #Array_S2, Cnt => #LEN_S2);
   #LEN := #LEN_S1 + #LEN_S2;
END_REGION

REGION Network 3
   #LWString_Connect := CONCAT(IN1 := #S1, IN2 := #S2);
END_REGION
END_FUNCTION

FUNCTION "Wchar_To_UTF8" : DWord   // FC162, SCL
{ S7_Optimized_Access := 'TRUE' }
VERSION : 0.1
   VAR_INPUT
      WChar : WChar;
   END_VAR
   VAR_OUTPUT
      Num : Int;
   END_VAR
   VAR_TEMP
      TempDword : DWord;
      Temp_Word : Word;
   END_VAR
BEGIN
   #Temp_Word := #WChar;
   #TempDword := W#16#0;
   IF 65535 > WORD_TO_UINT(#Temp_Word) AND WORD_TO_UINT(#Temp_Word)> 2048 THEN
       #TempDword.%X23 := 1;
       #TempDword.%X23 := 1;
       #TempDword.%X22 := 1;
       #TempDword.%X21 := 1;
       #TempDword.%X20 := 0;

       #TempDword.%X19 := #Temp_Word.%X15;
       #TempDword.%X18 := #Temp_Word.%X14;
       #TempDword.%X17 := #Temp_Word.%X13;
       #TempDword.%X16 := #Temp_Word.%X12;


       #TempDword.%X15 := 1;
       #TempDword.%X14 := 0;
       #TempDword.%X13 := #Temp_Word.%X11;
       #TempDword.%X12 := #Temp_Word.%X10;

       #TempDword.%X11 := #Temp_Word.%X9;
       #TempDword.%X10 := #Temp_Word.%X8;
       #TempDword.%X9 := #Temp_Word.%X7;
       #TempDword.%X8 := #Temp_Word.%X6;

       #TempDword.%X7 := 1;
       #TempDword.%X6 := 0;
       #TempDword.%X5 := #Temp_Word.%X5;
       #TempDword.%X4 := #Temp_Word.%X4;

       #TempDword.%X3 := #Temp_Word.%X3;
       #TempDword.%X2 := #Temp_Word.%X2;
       #TempDword.%X1 := #Temp_Word.%X1;
       #TempDword.%X0 := #Temp_Word.%X0;
       #Num := 3;


   ELSIF 2048 > WORD_TO_UINT(#Temp_Word) AND WORD_TO_UINT(#Temp_Word)> 128 THEN


       #TempDword.%X15 := 1;
       #TempDword.%X14 := 1;
       #TempDword.%X13 := 0;
       #TempDword.%X12 := #Temp_Word.%X10;

       #TempDword.%X11 := #Temp_Word.%X9;
       #TempDword.%X10 := #Temp_Word.%X8;
       #TempDword.%X9 := #Temp_Word.%X7;
       #TempDword.%X8 := #Temp_Word.%X6;

       #TempDword.%X7 := 1;
       #TempDword.%X6 := 0;
       #TempDword.%X5 := #Temp_Word.%X5;
       #TempDword.%X4 := #Temp_Word.%X4;

       #TempDword.%X3 := #Temp_Word.%X3;
       #TempDword.%X2 := #Temp_Word.%X2;
       #TempDword.%X1 := #Temp_Word.%X1;
       #TempDword.%X0 := #Temp_Word.%X0;
       #Num := 2;
   ELSE

       #TempDword.%X7 := 0;
       #TempDword.%X6 := #Temp_Word.%X6;
       #TempDword.%X5 := #Temp_Word.%X5;
       #TempDword.%X4 := #Temp_Word.%X4;

       #TempDword.%X3 := #Temp_Word.%X3;
       #TempDword.%X2 := #Temp_Word.%X2;
       #TempDword.%X1 := #Temp_Word.%X1;
       #TempDword.%X0 := #Temp_Word.%X0;
       #Num := 1;
   END_IF;
   #Wchar_To_UTF8 := #TempDword;
END_FUNCTION

// ===== library types =====

TYPE "HMI_SWD_Motor"
   STRUCT
      Start : Bool;
      Stop : Bool;
      REF : Real;
      TOR : Real;
      Ready : Bool;
      Running : Bool;
      Fault : Bool;
   END_STRUCT;
END_TYPE

TYPE "Step_By_Step"
   STRUCT
      StepNow : UInt;
      StepNum : UInt;
      StepName : String;
      StepReady : Bool;
      StepRuning : Bool;
      StepOK : Bool;
      StepNok : Bool;
   END_STRUCT;
END_TYPE

(* ===== HMI "HMI_RT_1" =====
system functions are stored by id; their names below are inferred from use
connection "HMI_连接_1": ETHERNET, S7_1200_OMS

HMI tags "默认变量表"
   "数据库字符串_Upload{11}" : 精炼机数据库 = PLC 数据库字符串.Upload[11], 1 s
   "数据库字符串_Upload{12}" : 精炼机数据库 = PLC 数据库字符串.Upload[12] AT %DB1.DBW0, 1 s
   "数据库字符串_Upload{13}" : 精炼机数据库 = PLC 数据库字符串.Upload[13] AT %DB1.DBW0, 1 s
   "数据库字符串_Upload{14}" : 精炼机数据库 = PLC 数据库字符串.Upload[14] AT %DB1.DBW0, 1 s
   "数据库字符串_Upload{15}" : 精炼机数据库 = PLC 数据库字符串.Upload[15] AT %DB1.DBW0, 1 s
   "通用数据采集_环境温度" : Real = PLC 通用数据采集.环境温度, 1 s
   "通用数据采集_环境湿度" : Real = PLC 通用数据采集.环境湿度, 1 s
   "精炼机数据转存_N21卷片机累计重量" : DInt = PLC 精炼机数据转存.N21卷片机累计重量 AT %DB100.DBD600, 1 s
   "精炼机数据转存_N22卷片机累计重量" : DInt = PLC 精炼机数据转存.N22卷片机累计重量 AT %DB100.DBD604, 1 s
   "数据库字符串_Query_Done" : Bool = PLC 数据库字符串.Query_Done, 1 s
   "数据库字符串_Connect_CND" : Bool = PLC 数据库字符串.Connect_CND, 1 s
   "数据库字符串_Query_Error" : Bool = PLC 数据库字符串.Query_Error, 1 s

HMI tags "系统变量"
   "Brightness" : Int, internal
   "ButtonDown" : Bool, internal
   "CodeView" : Bool, internal
   "CurrentLanguage" : Bool, internal
   "CurrentMachineState" : Int, internal
   "CurrentRecipeName" : WString[30], internal
   "CurrentUserName" : WString[18], internal
   "DiagState" : Int, internal
   "DummTagReal1" : LReal, internal
   "DummyDeltaInt" : Int, internal
   "DummyDeltaReal" : LReal, internal
   "DummyTagBool" : Bool, internal
   "DummyTagInt1" : Int, internal
   "DummyTagInt2" : Int, internal
   "DummyTagInt3" : Int, internal
   "InScreenTabState" : Int, internal
   "MainNavigationState" : Int, internal
   "OptionPanelNavigationState" : Int, internal
   "Password" : WString[20], internal
   "PopUpBackground" : Bool, internal
   "StartScreenName" : WString[60], internal
   "SubNavigationState" : Int, internal
   "ThirdLevelNavigationState" : Int, internal
   "TotalPieces" : Real, internal
   "UserIsLoggedIn" : Bool, internal
   "UserName" : WString[20], internal
   "InterAlarm" : Int, internal
   "EmergencyAuth" : Bool, internal
   "BM00_M001_Current_AlarmMax" : Real, internal
   "BM00_M001_Current_AlarmMin" : Real, internal
   "BM20_M001_Current_AlarmMax" : Real, internal
   "BM20_M001_Current_AlarmMin" : Real, internal

analog alarms
   1: '单螺杆过流报警', class Warnings, trigger "单螺杆电流滤波01_Ave"

text list "按钮名称": 0 'ON'; 1 'OFF'

text list "当前模式选择": 0 '演示模式'; 1 '测试模式'; 2 ''; 3 ''; 4 ''

text list "数据库状态": 0 '未连接'; 1 '已连接'; 2 '故障'

graphic list "DiagState_3": 0 'DiagOkay_White'; 1 'DiagWarning_White'; 2 'Circle'

screen "启动画面" 1920x1080, template "01_One_Nav_Level"
   GraphicView "图形视图_1" at 1,263 size 1608x666; Picture "rebuer_1"
   Button "按钮_1" at 1527,814 size 270x98; TextOff 'Entry'
      on Click: "MainEntry"()
   TextField "文本域_1" at 626,494 size 773x90; Text '江苏睿博环保设备有限公司'
   TextField "文本域_2" at 630,580 size 676x68; Text 'REB-ZSI型智能废橡胶精炼设备'